HMI tags "DB_SDC_EMS"
   "SDC\DB_SDC_EMS\EMS[XXX].DISTANCE" : DInt AT %DB0.DBD0, 1 s   // Abstand zum vorangehenden EMS / distance to preciding EMS
   "SDC\DB_SDC_EMS\_Byte_EMS[XXX].ABS_POS" : Int, internal   // Absolute Position / absolute Positon
   "SDC\DB_SDC_EMS\EMS[XXX].IF_I_EMS.STAT" : DWord AT %DB0.DBD0, 1 s
   "SDC\DB_SDC_EMS\EMS[XXX].PRECEDING_EMS" : Int AT %DB0.DBW0, 1 s   // preciding EMS
   "SDC\DB_SDC_EMS\_Byte_EMS[XXX].TS_STAT.VAL.SEK" : Int, internal   // Sektion
   "SDC\DB_SDC_EMS\_Byte_EMS[XXX].DISTANCE" : Int, internal   // Abstand zum vorangehenden EMS / distance to preciding EMS
   "DB_SDC_EMS_HMI_HEADER.START_HMI" : Int = PLC DB_SDC_EMS_HMI.HEADER.START_HMI AT %DB3814.DBW16, 1 s   // Startadresse HMI
   "SDC\DB_SDC_EMS\EMS[XXX].IF_I_EMS.EA1" : DWord AT %DB0.DBD0, 1 s
   "SDC\DB_SDC_EMS\HMI[XX].PROFIL_Nr" : Int AT %DB0.DBW0, 1 s   // Profilnummer
   "SDC\DB_SDC_EMS\_EMS_HMI_Byte_16" : Int, internal
   "SDC\DB_SDC_EMS\HMI[XX].T_EDIT" : Bool AT %DB0.DBX0.0, 1 s   // Taster Editieren für Pult aktivieren
   "SDC\DB_SDC_EMS\_EMS_HMI_Byte_18" : Int, internal
   "SDC\DB_SDC_EMS\EMS[XXX].FKT_RESET" : Word AT %DB0.DBW0, 1 s   // EMS zur Reperatur / EMS to Repair
   "SDC\DB_SDC_EMS\EMS[XXX].IF_Q_EMS.D_SETSPEED" : DInt AT %DB0.DBD0, 1 s   // set value: drive speed (mm/min)
   "SDC\DB_SDC_EMS\_Byte_EMS[XXX].CYCLE_COUNTER" : Int, internal   // Zykluszähler / Cycle Counter
   "SDC\DB_SDC_EMS\HMI[XX].FR_EDIT" : Bool AT %DB0.DBX0.0, 1 s   // Freigabe Editieren
   "SDC\DB_SDC_EMS\_Byte_EMS[XXX].IF_I_EMS.H_POS" : Int, internal
   "SDC\DB_SDC_EMS\EMS[XXX].TS_STAT.SERIES" : Array [0..3] of Char AT %DB0.DBX0.0, 1 s   // Entwicklungs Serie Karosse (e.g. E-90, E-87 ) / Development series body (e.g. E-90, E-87 )
   "SDC\DB_SDC_EMS\EMS[XXX].IF_Q_EMS.D_SETPOS" : DInt AT %DB0.DBD0, 1 s   // Setpoint: drive position in mm
   "SDC\DB_SDC_EMS\HMI[XX].BILD_Nr_Alt" : Int AT %DB0.DBW0, 1 s   // Bild_Nr alt
   "SDC\DB_SDC_EMS\EMS[XXX].IF_Q_EMS.H_SETSPEED" : Int AT %DB0.DBW0, 1 s   // Setpoint: hoist speed (mm/min)
   "SDC\DB_SDC_EMS\_EMS_HMI_Byte_10" : Int, internal
   "SDC\DB_SDC_EMS\EMS[XXX].IF_I_EMS.H_POS" : Int AT %DB0.DBW0, 1 s
   "SDC\DB_SDC_EMS\_Byte_EMS[XXX].IF_Q_EMS.D_SETPOS" : Int, internal   // Setpoint: drive position in mm Pointer
   "SDC\DB_SDC_EMS\HMI[XX].EMS_Nr" : Int AT %DB0.DBW0, 1 s   // Sektionsnummer
   "SDC\DB_SDC_EMS\_Byte_EMS[XXX].PRECEDING_EMS" : Int, internal   // preciding EMS
   "SDC\DB_SDC_EMS\_Byte_EMS[XXX].IF_I_EMS.STAT" : Int, internal
   "SDC\DB_SDC_EMS\_EMS_HMI_Byte_09" : Int, internal
   "SDC\DB_SDC_EMS\_Byte_EMS[XXX].ERRORS_SDC" : Int, internal   // Fehler SDC Pointer / Faults SDC Pointer
   "SDC\DB_SDC_EMS\EMS[XXX].FLAGS" : Word AT %DB0.DBW0, 1 s   // EMS antrieb vorhanden / EMSdriver present
   "SDC\DB_SDC_EMS\_Byte_EMS[XXX].IF_I_EMS.EA2" : Int, internal
   "SDC\DB_SDC_EMS\EMS[XXX].ERRORS_SDC" : Word AT %DB0.DBW0, 1 s   // Fehler SDC / Faults SDC
   "SDC\DB_SDC_EMS\HMI[XX].T_SAVE" : Bool AT %DB0.DBX0.2, 1 s   // Taster speichern
   "SDC\DB_SDC_EMS\_Byte_EMS[XXX].PROFIL" : Int, internal   // Profile Number
   "SDC\DB_SDC_EMS\_Byte_EMS[XXX].FLAGS" : Int, internal   // EMS antrieb vorhanden / EMSdriver present
   "DB_SDC_EMS_1_HEADER.START_EMS" : Int = PLC DB_SDC_EMS_1.HEADER.START_EMS AT %DB3714.DBW6, 1 s   // Startadresse der EMS Daten im Daten DB
   "SDC\DB_SDC_EMS\EMS[XXX].IF_I_EMS.EA2" : DWord AT %DB0.DBD0, 1 s
   "SDC\DB_SDC_EMS\EMS[XXX].TS_STAT.VAL.SEK" : Int AT %DB0.DBW0, 1 s   // Sektion
      on ChangeValue: "SDC_TS_REFERENCE"("SDC\DB_SDC_EMS\EMS[XXX].TS_STAT.VAL.SEK")
   "SDC\DB_SDC_EMS\EMS[XXX].IF_I_EMS.D_POS" : DInt AT %DB0.DBD0, 1 s
   "SDC\DB_SDC_EMS\_Byte_EMS[XXX].IF_Q_EMS.H_SETSPEED" : Int, internal   // Setpoint: hoist speed (mm/min) Pointer
   "DB_SDC_EMS_1_HEADER.LAENGE_EMS" : Int = PLC DB_SDC_EMS_1.HEADER.LAENGE_EMS AT %DB3714.DBW8, 1 s   // Länge Eingänge pro EMS
   "SDC\DB_SDC_EMS\_EMS_HMI_Byte_19" : Int, internal
   "DB_SDC_EMS_1_HEADER.MIN_NR_EMS" : Int = PLC DB_SDC_EMS_1.HEADER.MIN_NR_EMS AT %DB3714.DBW2, 1 s   // Niedrigste EMS Nummer im Daten DB
   "SDC\DB_SDC_EMS\_Byte_EMS[XXX].IF_Q_EMS.H_SETPOS" : Int, internal   // Setpoint: hoist position (mm) Pointer
   "SDC\DB_SDC_EMS\_Byte_EMS[XXX].IF_I_EMS.EA1" : Int, internal
   "SDC\DB_SDC_EMS\_Intern_DB_EMS_Nr" : Int, internal
   "SDC\DB_SDC_EMS\HMI[XX].ER_DATA" : Bool AT %DB0.DBX0.1, 1 s   // Daten Fehlerhaft
   "DB_SDC_EMS_1_HEADER.OFFSET_EMS_FKT" : Int = PLC DB_SDC_EMS_1.HEADER.OFFSET_EMS_FKT AT %DB3714.DBW14, 1 s   // Offset EMS Funktions
   "SDC\DB_SDC_EMS\EMS[XXX].IF_Q_EMS.H_SETPOS" : Int AT %DB0.DBW0, 1 s   // Setpoint: hoist position (mm)
   "SDC\DB_SDC_EMS\_Byte_EMS[XXX].IF_I_EMS.ERROR" : Int, internal   // Fehlernummer Pointer / Error number Pointer
   "SDC\DB_SDC_EMS\_Byte_EMS[XXX].FKT_RESET" : Int, internal   // EMS zur Reperatur / EMS to Repair
   "SDC\DB_SDC_EMS\EMS[XXX].IF_Q_EMS.CONT" : DWord AT %DB0.DBD0, 1 s
   "DB_SDC_EMS_HMI_HEADER.OFFEST_HMI_DATA" : Int = PLC DB_SDC_EMS_HMI.HEADER.OFFEST_HMI_DATA AT %DB3814.DBW18, 1 s   // Offestadresse der HMI EMS Data
   "SDC\DB_SDC_EMS\_Byte_EMS[XXX].FKT_SET" : Int, internal   // EMS zur Reperatur / EMS to Repair
   "SDC\DB_SDC_EMS\HMI[XX].PULT_Nr_EDIT" : Int AT %DB0.DBW0, 1 s   // Pult Nr Editieren Aktiv (HMI 1 = Master)
   "SDC\DB_SDC_EMS\_EMS_HMI_Byte_00" : Int, internal
   "DB_SDC_EMS_1_HEADER.MAX_NR_EMS" : Int = PLC DB_SDC_EMS_1.HEADER.MAX_NR_EMS AT %DB3714.DBW4, 1 s   // Höchste EMS Nummer im Daten DB
   "SDC\DB_SDC_EMS\EMS[XXX].IF_I_EMS.ERROR" : Int AT %DB0.DBW0, 1 s   // Fehlernummer / Error number
   "DB_SDC_EMS_1_HEADER.OFFSET_EMS_SEK_STAT" : Int = PLC DB_SDC_EMS_1.HEADER.OFFSET_EMS_SEK_STAT AT %DB3714.DBW10, 1 s   // Offset EMS Data
   "DB_SDC_EMS_1_HEADER.LAENGE_EMS_SEK_STAT" : Int = PLC DB_SDC_EMS_1.HEADER.LAENGE_EMS_SEK_STAT AT %DB3714.DBW12, 1 s   // Länge EMS Data
   "SDC\DB_SDC_EMS\_Byte_EMS[XXX].TS_STAT.SERIES" : Int, internal   // Entwicklungs Serie Karosse (e.g. E-90, E-87 ) / Development series body (e.g. E-90, E-87 )
   "SDC\DB_SDC_EMS\HMI[XX].BILD_Nr" : Int AT %DB0.DBW0, 1 s   // Bild_Nr aktiv
   "SDC\DB_SDC_EMS\EMS[XXX].CYCLE_COUNTER" : Int AT %DB0.DBW0, 1 s   // Zykluszähler / Cycle Counter
   "SDC\DB_SDC_EMS\EMS[XXX].FKT_SET" : Word AT %DB0.DBW0, 1 s   // EMS zur Reperatur / EMS to Repair
      on ChangeValue: ResetBit("SDC\DB_SDC_EMS\_Intern_EMS_FKT_Info_Rep_1_on"); ResetBit("SDC\DB_SDC_EMS\_Intern_EMS_FKT_Info_Rep_2_on")
   "SDC\DB_SDC_EMS\HMI[XX].T_LOAD" : Bool AT %DB0.DBX0.3, 1 s   // Taster laden
   "SDC\DB_SDC_EMS\_EMS_HMI_Byte_12" : Int, internal
   "SDC\DB_SDC_EMS\_EMS_HMI_Byte_04" : Int, internal
   "DB_SDC_EMS_HMI_HMI[1].PULT_Nr_EDIT" : Int = PLC DB_SDC_EMS_HMI.HMI[1].PULT_Nr_EDIT AT %DB3814.DBW20, 1 s   // Pult Nr Editieren Aktiv (HMI 1 = Master)
   "SDC\DB_SDC_EMS\_EMS_HMI_Byte_14" : Int, internal
   "SDC\DB_SDC_EMS\_EMS_HMI_Byte_06" : Int, internal
   "SDC\DB_SDC_EMS\_Byte_EMS[XXX].IF_I_EMS.D_POS" : Int, internal
   "SDC\DB_SDC_EMS\_EMS_HMI_Byte_08" : Int, internal
   "SDC\DB_SDC_EMS\EMS[XXX].PROFIL" : Int AT %DB0.DBW0, 1 s   // Profile Number
      on ChangeValue: "SDC_GLOBAL_REFERENCE_PROFIL"("SDC\DB_SDC_EMS\EMS[XXX].PROFIL")
   "SDC\DB_SDC_EMS\_EMS_HMI_Byte_02" : Int, internal
   "SDC\DB_SDC_EMS\EMS[XXX].ABS_POS" : DInt AT %DB0.DBD0, 1 s   // absolute Positon
   "SDC\DB_SDC_EMS\HMI[XX].T_RESET_BED" : Bool AT %DB0.DBX0.1, 1 s   // Taster Reset Bedienfreigabe Pult Nr Bedienung
   "SDC\DB_SDC_EMS\_Byte_EMS[XXX].IF_Q_EMS.CONT" : Int, internal
   "SDC\DB_SDC_EMS\_Byte_EMS[XXX].IF_Q_EMS.D_SETSPEED" : Int, internal   // set value: drive speed (mm/min) Pointer
   "SDC\DB_SDC_EMS\_Byte_EMS[XXX].TS_STAT.VAL.ERROR" : Int, internal   // Sektion
   "SDC\DB_SDC_EMS\EMS[XXX].TS_STAT.VAL.ERROR" : Int AT %DB0.DBW0, 1 s   // Sektion
      on ChangeValue: SetTag("_DB_SDC_ERRORS.Error_nr", "SDC\DB_SDC_EMS\EMS[XXX].TS_STAT.VAL.ERROR")
   "DB_SDC_EMS_HMI_HEADER.DB_NR" : Int = PLC DB_SDC_EMS_HMI.HEADER.DB_NR AT %DB3814.DBW0, 1 s   // DB Nummer
   "SDC\DB_SDC_EMS\_Byte_EMS[XXX].IF_Q_EMS.T_SETPOS" : Int, internal   // Setpoint: hoist position (mm) Pointer
   "SDC\DB_SDC_EMS\_Byte_EMS[XXX].IF_Q_EMS.T_SETSPEED" : Int, internal   // Setpoint: hoist speed (mm/min) Pointer
   "SDC\DB_SDC_EMS\EMS[XXX].IF_Q_EMS.T_SETPOS" : Int AT %DB0.DBW0, 1 s   // Setpoint: hoist position (mm)
   "SDC\DB_SDC_EMS\EMS[XXX].IF_Q_EMS.T_SETSPEED" : Int AT %DB0.DBW0, 1 s   // Setpoint: hoist speed (mm/min)
   "SDC\DB_SDC_EMS\_Byte_EMS[XXX].IF_I_EMS.T_POS" : Int, internal
   "SDC\DB_SDC_EMS\EMS[XXX].IF_I_EMS.T_POS" : Int AT %DB0.DBW0, 1 s
   "SDC\DB_SDC_EMS\_Byte_EMS[XXX].FKT_INFO_REP_1" : Int, internal
   "SDC\DB_SDC_EMS\_Byte_EMS[XXX].FKT_INFO_REP_2" : Int, internal
   "SDC\DB_SDC_EMS\EMS[XXX].FKT_INFO_REP_1" : Int AT %DB0.DBW0, 1 s
   "SDC\DB_SDC_EMS\EMS[XXX].FKT_INFO_REP_2" : Int AT %DB0.DBW0, 1 s
   "SDC\DB_SDC_EMS\_Intern_EMS_FKT_Info_Rep_1_on" : Bool, internal
   "SDC\DB_SDC_EMS\_Intern_EMS_FKT_Info_Rep_2_on" : Bool, internal
   "SDC\DB_SDC_EMS\EMS[XXX].IF_I_EMS.EA3" : Word AT %DB0.DBW0, 1 s
   "SDC\DB_SDC_EMS\_Byte_EMS[XXX].IF_I_EMS.EA3" : Int, internal
   "SDC\DB_SDC_EMS\_Byte_EMS[XXX].VersNo[0]" : Int, internal   // Zykluszähler / Cycle Counter
   "SDC\DB_SDC_EMS\_Byte_EMS[XXX].VersNo[1]" : Int, internal   // Zykluszähler / Cycle Counter
   "SDC\DB_SDC_EMS\EMS[XXX].VersNo[0]" : Byte AT %DB0.DBB0, 1 s   // Zykluszähler / Cycle Counter
   "SDC\DB_SDC_EMS\EMS[XXX].VersNo[1]" : Byte AT %DB0.DBB0, 1 s   // Zykluszähler / Cycle Counter

HMI tags "DB_SDC_SIM"
   "DB_SDC_EMS_SIM_PAR.ON" : Bool = PLC DB_SDC_EMS_SIM.PAR.ON AT %DB3726.DBX40.0, 1 s   // Simulation ON "1"
   "DB_SDC_EMS_SIM_PAR.LEAP_AKT" : Array [0..19] of Bool = PLC DB_SDC_EMS_SIM.PAR.LEAP_AKT AT %DB3726.DBX32.0, 1 s   // Leap Aktiv
   "DB_SDC_EMS_SIM_PAR.BARCODE_START" : DInt = PLC DB_SDC_EMS_SIM.PAR.BARCODE_START AT %DB3726.DBD20, 1 s   // min Barcodevalue
   "DB_SDC_EMS_SIM_PAR.HUB_ENDE" : Int = PLC DB_SDC_EMS_SIM.PAR.HUB_ENDE AT %DB3726.DBW30, 1 s   // max Hoistvalue
   "DB_SDC_EMS_SIM_EMS[2].D_POS" : DInt = PLC DB_SDC_EMS_SIM.EMS[2].D_POS AT %DB3726.DBD90, 1 s   // Antriebsposition in mm / Drive position in mm
   "DB_SDC_EMS_SIM_PAR.BARCODE_ENDE" : DInt = PLC DB_SDC_EMS_SIM.PAR.BARCODE_ENDE AT %DB3726.DBD24, 1 s   // max Barcodevalue
   "DB_SDC_EMS_SIM_PAR.HUB_START" : Int = PLC DB_SDC_EMS_SIM.PAR.HUB_START AT %DB3726.DBW28, 1 s   // min Hoistvalue
   "DB_SDC_EMS_SIM_EMS[1].D_POS" : DInt = PLC DB_SDC_EMS_SIM.EMS[1].D_POS AT %DB3726.DBD50, 1 s   // Antriebsposition in mm / Drive position in mm
   "DB_SDC_EMS_SIM_EMS[3].D_POS" : DInt = PLC DB_SDC_EMS_SIM.EMS[3].D_POS AT %DB3726.DBD130, 1 s   // Antriebsposition in mm / Drive position in mm

HMI tags "DB_SDC_ERRORS"
   "DB_SDC_ERRORS_HEADER.DB_NR" : Int = PLC DB_SDC_ERRORS.HEADER.DB_NR AT %DB3722.DBW0, 1 s
   "DB_SDC_ERRORS_HEADER.MIN_NR_EMS" : Int = PLC DB_SDC_ERRORS.HEADER.MIN_NR_EMS AT %DB3722.DBW2, 1 s
   "DB_SDC_ERRORS_HEADER.MAX_NR_EMS" : Int = PLC DB_SDC_ERRORS.HEADER.MAX_NR_EMS AT %DB3722.DBW4, 1 s
   "DB_SDC_ERRORS_HEADER.START_EMS" : Int = PLC DB_SDC_ERRORS.HEADER.START_EMS AT %DB3722.DBW6, 1 s
   "DB_SDC_ERRORS_HEADER.LAENGE_EMS_StörungS" : Int = PLC DB_SDC_ERRORS.HEADER.LAENGE_EMS_StörungS AT %DB3722.DBW8, 1 s
   "DB_SDC_ERRORS.EMS[XXX].GEN_1" : Word AT %DB0.DBW0, 1 s
   "_Byte_DB_SDC_ERRORS.EMS[XXX].GEN_1" : UInt, internal
   "DB_SDC_ERRORS.EMS[XXX].GEN_2" : Word AT %DB0.DBW0, 1 s
   "_Byte_DB_SDC_ERRORS.EMS[XXX].GEN_2" : UInt, internal
   "DB_SDC_ERRORS.EMS[XXX].GEN_3" : Word AT %DB0.DBW0, 1 s
   "_Byte_DB_SDC_ERRORS.EMS[XXX].GEN_3" : UInt, internal
   "DB_SDC_ERRORS.EMS[XXX].GEN_4" : Word AT %DB0.DBW0, 1 s
   "_Byte_DB_SDC_ERRORS.EMS[XXX].GEN_4" : UInt, internal
   "DB_SDC_ERRORS.EMS[XXX].DRIVE_1" : Word AT %DB0.DBW0, 1 s
   "_Byte_DB_SDC_ERRORS.EMS[XXX].DRIVE_1" : UInt, internal
   "DB_SDC_ERRORS.EMS[XXX].DRIVE_2" : Word AT %DB0.DBW0, 1 s
   "_Byte_DB_SDC_ERRORS.EMS[XXX].DRIVE_2" : UInt, internal
   "DB_SDC_ERRORS.EMS[XXX].FC_DRIVE_1" : Word AT %DB0.DBW0, 1 s
   "_Byte_DB_SDC_ERRORS.EMS[XXX].FC_DRIVE_1" : UInt, internal
   "DB_SDC_ERRORS.EMS[XXX].FC_DRIVE_2" : Word AT %DB0.DBW0, 1 s
   "_Byte_DB_SDC_ERRORS.EMS[XXX].FC_DRIVE_2" : UInt, internal
   "DB_SDC_ERRORS.EMS[XXX].SAFETY_DRIVE" : Word AT %DB0.DBW0, 1 s
   "_Byte_DB_SDC_ERRORS.EMS[XXX].SAFETY_DRIVE" : UInt, internal
   "_Byte_DB_SDC_ERRORS.EMS[XXX].HOIST_1" : UInt, internal
   "DB_SDC_ERRORS.EMS[XXX].HOIST_2" : Word AT %DB0.DBW0, 1 s
   "_Byte_DB_SDC_ERRORS.EMS[XXX].HOIST_2" : UInt, internal
   "DB_SDC_ERRORS.EMS[XXX].FC_HOIST_1" : Word AT %DB0.DBW0, 1 s
   "_Byte_DB_SDC_ERRORS.EMS[XXX].FC_HOIST_1" : UInt, internal
   "DB_SDC_ERRORS.EMS[XXX].FC_HOIST_2" : Word AT %DB0.DBW0, 1 s
   "_Byte_DB_SDC_ERRORS.EMS[XXX].FC_HOIST_2" : UInt, internal
   "DB_SDC_ERRORS.EMS[XXX].SAFETY_HOIST" : Word AT %DB0.DBW0, 1 s
   "_Byte_DB_SDC_ERRORS.EMS[XXX].SAFETY_HOIST" : UInt, internal
   "DB_SDC_ERRORS.EMS[XXX].HOIST_1" : Word AT %DB0.DBW0, 1 s
   "_Byte_DB_SDC_ERRORS.EMS[XXX].TILT_1" : UInt, internal
   "DB_SDC_ERRORS.EMS[XXX].TILT_2" : Word AT %DB0.DBW0, 1 s
   "_Byte_DB_SDC_ERRORS.EMS[XXX].TILT_2" : UInt, internal
   "DB_SDC_ERRORS.EMS[XXX].FC_TILT_1" : Word AT %DB0.DBW0, 1 s
   "_Byte_DB_SDC_ERRORS.EMS[XXX].FC_TILT_1" : UInt, internal
   "DB_SDC_ERRORS.EMS[XXX].FC_TILT_2" : Word AT %DB0.DBW0, 1 s
   "_Byte_DB_SDC_ERRORS.EMS[XXX].FC_TILT_2" : UInt, internal
   "DB_SDC_ERRORS.EMS[XXX].SAFETY_TILT" : Word AT %DB0.DBW0, 1 s
   "_Byte_DB_SDC_ERRORS.EMS[XXX].SAFETY_TILT" : UInt, internal
   "DB_SDC_ERRORS.EMS[XXX].TILT_1" : Word AT %DB0.DBW0, 1 s
   "DB_SDC_ERRORS.EMS[XXX].SDC" : Word AT %DB0.DBW0, 1 s
   "_Byte_DB_SDC_ERRORS.EMS[XXX].SDC" : UInt, internal
   "DB_SDC_ERRORS.SDC" : Word AT %DB3722.DBW20020, 1 s
   "_DB_SDC_ERRORS.Error_nr" : Int, internal

HMI tags "DB_SDC_GLOBAL_REFERENCE"
   "DB_SDC_GLOBAL_REFERENCE_PAR_SET[8].LIMITS" : Array [0..15] of Char = PLC DB_SDC_GLOBAL_REFERENCE.PAR_SET[8].LIMITS AT %DB3786.DBX292.0, 1 s
   "DB_SDC_GLOBAL_REFERENCE_PAR_SET[3].LIMITS" : Array [0..15] of Char = PLC DB_SDC_GLOBAL_REFERENCE.PAR_SET[3].LIMITS AT %DB3786.DBX132.0, 1 s
   "DB_SDC_GLOBAL_REFERENCE_PAR_SET[0].LIMITS" : Array [0..15] of Char = PLC DB_SDC_GLOBAL_REFERENCE.PAR_SET[0].LIMITS AT %DB3786.DBX36.0, 1 s
   "DB_SDC_GLOBAL_REFERENCE_PAR_SET[14].SYNCH" : Array [0..15] of Char = PLC DB_SDC_GLOBAL_REFERENCE.PAR_SET[14].SYNCH AT %DB3786.DBX468.0, 1 s
   "DB_SDC_GLOBAL_REFERENCE_PAR_SET[9].SYNCH" : Array [0..15] of Char = PLC DB_SDC_GLOBAL_REFERENCE.PAR_SET[9].SYNCH AT %DB3786.DBX308.0, 1 s
   "DB_SDC_GLOBAL_REFERENCE_PAR_SET[11].LIMITS" : Array [0..15] of Char = PLC DB_SDC_GLOBAL_REFERENCE.PAR_SET[11].LIMITS AT %DB3786.DBX388.0, 1 s
   "DB_SDC_GLOBAL_REFERENCE_PAR_SET[10].LIMITS" : Array [0..15] of Char = PLC DB_SDC_GLOBAL_REFERENCE.PAR_SET[10].LIMITS AT %DB3786.DBX356.0, 1 s
   "DB_SDC_GLOBAL_REFERENCE_PAR_SET[0].SYNCH" : Array [0..15] of Char = PLC DB_SDC_GLOBAL_REFERENCE.PAR_SET[0].SYNCH AT %DB3786.DBX20.0, 1 s
   "DB_SDC_GLOBAL_REFERENCE_PAR_SET[14].LIMITS" : Array [0..15] of Char = PLC DB_SDC_GLOBAL_REFERENCE.PAR_SET[14].LIMITS AT %DB3786.DBX484.0, 1 s
   "DB_SDC_GLOBAL_REFERENCE_PAR_SET[6].LIMITS" : Array [0..15] of Char = PLC DB_SDC_GLOBAL_REFERENCE.PAR_SET[6].LIMITS AT %DB3786.DBX228.0, 1 s
   "DB_SDC_GLOBAL_REFERENCE_PAR_SET[10].SYNCH" : Array [0..15] of Char = PLC DB_SDC_GLOBAL_REFERENCE.PAR_SET[10].SYNCH AT %DB3786.DBX340.0, 1 s
   "DB_SDC_GLOBAL_REFERENCE_PAR_SET[5].SYNCH" : Array [0..15] of Char = PLC DB_SDC_GLOBAL_REFERENCE.PAR_SET[5].SYNCH AT %DB3786.DBX180.0, 1 s
   "DB_SDC_GLOBAL_REFERENCE_PAR_SET[13].SYNCH" : Array [0..15] of Char = PLC DB_SDC_GLOBAL_REFERENCE.PAR_SET[13].SYNCH AT %DB3786.DBX436.0, 1 s
   "DB_SDC_GLOBAL_REFERENCE_PAR_SET[12].LIMITS" : Array [0..15] of Char = PLC DB_SDC_GLOBAL_REFERENCE.PAR_SET[12].LIMITS AT %DB3786.DBX420.0, 1 s
   "DB_SDC_GLOBAL_REFERENCE_PAR_SET[15].SYNCH" : Array [0..15] of Char = PLC DB_SDC_GLOBAL_REFERENCE.PAR_SET[15].SYNCH AT %DB3786.DBX500.0, 1 s
   "DB_SDC_GLOBAL_REFERENCE_PAR_SET[2].LIMITS" : Array [0..15] of Char = PLC DB_SDC_GLOBAL_REFERENCE.PAR_SET[2].LIMITS AT %DB3786.DBX100.0, 1 s
   "DB_SDC_GLOBAL_REFERENCE_PAR_SET[6].SYNCH" : Array [0..15] of Char = PLC DB_SDC_GLOBAL_REFERENCE.PAR_SET[6].SYNCH AT %DB3786.DBX212.0, 1 s
   "DB_SDC_GLOBAL_REFERENCE_PAR_SET[1].SYNCH" : Array [0..15] of Char = PLC DB_SDC_GLOBAL_REFERENCE.PAR_SET[1].SYNCH AT %DB3786.DBX52.0, 1 s
   "DB_SDC_GLOBAL_REFERENCE_PAR_SET[4].SYNCH" : Array [0..15] of Char = PLC DB_SDC_GLOBAL_REFERENCE.PAR_SET[4].SYNCH AT %DB3786.DBX148.0, 1 s
   "DB_SDC_GLOBAL_REFERENCE_PAR_SET[8].SYNCH" : Array [0..15] of Char = PLC DB_SDC_GLOBAL_REFERENCE.PAR_SET[8].SYNCH AT %DB3786.DBX276.0, 1 s
   "DB_SDC_GLOBAL_REFERENCE_PAR_SET[2].SYNCH" : Array [0..15] of Char = PLC DB_SDC_GLOBAL_REFERENCE.PAR_SET[2].SYNCH AT %DB3786.DBX84.0, 1 s
   "DB_SDC_GLOBAL_REFERENCE_PAR_SET[1].LIMITS" : Array [0..15] of Char = PLC DB_SDC_GLOBAL_REFERENCE.PAR_SET[1].LIMITS AT %DB3786.DBX68.0, 1 s
   "DB_SDC_GLOBAL_REFERENCE_PAR_SET[15].LIMITS" : Array [0..15] of Char = PLC DB_SDC_GLOBAL_REFERENCE.PAR_SET[15].LIMITS AT %DB3786.DBX516.0, 1 s
   "DB_SDC_GLOBAL_REFERENCE_PAR_SET[11].SYNCH" : Array [0..15] of Char = PLC DB_SDC_GLOBAL_REFERENCE.PAR_SET[11].SYNCH AT %DB3786.DBX372.0, 1 s
   "DB_SDC_GLOBAL_REFERENCE_PAR_SET[3].SYNCH" : Array [0..15] of Char = PLC DB_SDC_GLOBAL_REFERENCE.PAR_SET[3].SYNCH AT %DB3786.DBX116.0, 1 s
   "DB_SDC_GLOBAL_REFERENCE_PAR_SET[4].LIMITS" : Array [0..15] of Char = PLC DB_SDC_GLOBAL_REFERENCE.PAR_SET[4].LIMITS AT %DB3786.DBX164.0, 1 s
   "DB_SDC_GLOBAL_REFERENCE_PAR_SET[12].SYNCH" : Array [0..15] of Char = PLC DB_SDC_GLOBAL_REFERENCE.PAR_SET[12].SYNCH AT %DB3786.DBX404.0, 1 s
   "DB_SDC_GLOBAL_REFERENCE_PAR_SET[9].LIMITS" : Array [0..15] of Char = PLC DB_SDC_GLOBAL_REFERENCE.PAR_SET[9].LIMITS AT %DB3786.DBX324.0, 1 s
   "DB_SDC_GLOBAL_REFERENCE_PAR_SET[7].SYNCH" : Array [0..15] of Char = PLC DB_SDC_GLOBAL_REFERENCE.PAR_SET[7].SYNCH AT %DB3786.DBX244.0, 1 s
   "DB_SDC_GLOBAL_REFERENCE_PAR_SET[7].LIMITS" : Array [0..15] of Char = PLC DB_SDC_GLOBAL_REFERENCE.PAR_SET[7].LIMITS AT %DB3786.DBX260.0, 1 s
   "DB_SDC_GLOBAL_REFERENCE_PAR_SET[13].LIMITS" : Array [0..15] of Char = PLC DB_SDC_GLOBAL_REFERENCE.PAR_SET[13].LIMITS AT %DB3786.DBX452.0, 1 s
   "DB_SDC_GLOBAL_REFERENCE_PAR_SET[5].LIMITS" : Array [0..15] of Char = PLC DB_SDC_GLOBAL_REFERENCE.PAR_SET[5].LIMITS AT %DB3786.DBX196.0, 1 s
   "SDC\DB_SDC_GLOBAL_REFERENCE\DB_SDC_GLOBAL_REFERENCE.PROFIL[XX].SORTE" : Array [0..5] of Char AT %DB0.DBX0.0, 1 s
   "DB_SDC_GLOBAL_REFERENCE_HEADER.START_PROFIL" : Int = PLC DB_SDC_GLOBAL_REFERENCE.HEADER.START_PROFIL AT %DB3786.DBW14, 1 s
   "DB_SDC_GLOBAL_REFERENCE_HEADER.LAENGE_PROFIL" : Int = PLC DB_SDC_GLOBAL_REFERENCE.HEADER.LAENGE_PROFIL AT %DB3786.DBW16, 1 s
   "_DB_SDC_GLOBAL_REFERENCE.PROFIL[XX].SORTE_Byte" : Int, internal
   "DB_SDC_GLOBAL_REFERENCE_HEADER.MIN_PROFIL" : Int = PLC DB_SDC_GLOBAL_REFERENCE.HEADER.MIN_PROFIL AT %DB3786.DBW10, 1 s
   "DB_SDC_GLOBAL_REFERENCE_HEADER.MAX_PROFIL" : Int = PLC DB_SDC_GLOBAL_REFERENCE.HEADER.MAX_PROFIL AT %DB3786.DBW12, 1 s
   "_DB_SDC_GLOBAL_REFERENCE.PROFIL[XX+1].SORTE_Byte" : Int, internal
   "SDC\DB_SDC_GLOBAL_REFERENCE\DB_SDC_GLOBAL_REFERENCE.PROFIL[XX+1].SORTE" : Array [0..5] of Char AT %DB0.DBX0.0, 1 s
   "DB_SDC_GLOBAL_REFERENCE_HEADER.DB_NR" : Int = PLC DB_SDC_GLOBAL_REFERENCE.HEADER.DB_NR AT %DB3786.DBW0, 1 s

HMI tags "DB_SDC_EMS_TA"
   "DB_SDC_EMS_TA_HEADER.DB_NR" : Int = PLC DB_SDC_EMS_TA.HEADER.DB_NR AT %DB3728.DBW0, 1 s
   "DB_SDC_EMS_TA_HEADER.MIN_NR_EMS" : Int = PLC DB_SDC_EMS_TA.HEADER.MIN_NR_EMS AT %DB3728.DBW2, 1 s
   "DB_SDC_EMS_TA_HEADER.MAX_NR_EMS" : Int = PLC DB_SDC_EMS_TA.HEADER.MAX_NR_EMS AT %DB3728.DBW4, 1 s
   "DB_SDC_EMS_TA_HEADER.START_EMS" : Int = PLC DB_SDC_EMS_TA.HEADER.START_EMS AT %DB3728.DBW6, 1 s
   "DB_SDC_EMS_TA_HEADER.LAENGE_TA_DATA" : Int = PLC DB_SDC_EMS_TA.HEADER.LAENGE_TA_DATA AT %DB3728.DBW8, 1 s
   "DB_SDC_EMS_TA_HEADER.ANZ_TA" : Int = PLC DB_SDC_EMS_TA.HEADER.ANZ_TA AT %DB3728.DBW10, 1 s
   "DB_SDC_EMS_TA.EMS[XX].TA1.PW1" : Int AT %DB0.DBW0, 1 s
   "_Byte_DB_SDC_EMS_TA.EMS[XX].TA1.PW1" : DInt, internal
   "_Byte_DB_SDC_EMS_TA.EMS[XX].TA1.PW2" : DInt, internal
   "_Byte_DB_SDC_EMS_TA.EMS[XX].TA1.PW3" : DInt, internal
   "_Byte_DB_SDC_EMS_TA.EMS[XX].TA2.PW1" : DInt, internal
   "_Byte_DB_SDC_EMS_TA.EMS[XX].TA2.PW2" : DInt, internal
   "_Byte_DB_SDC_EMS_TA.EMS[XX].TA2.PW3" : DInt, internal
   "_Byte_DB_SDC_EMS_TA.EMS[XX].TA3.PW1" : DInt, internal
   "_Byte_DB_SDC_EMS_TA.EMS[XX].TA3.PW2" : DInt, internal
   "_Byte_DB_SDC_EMS_TA.EMS[XX].TA3.PW3" : DInt, internal
   "DB_SDC_EMS_TA.EMS[XX].TA1.PW2" : Int AT %DB0.DBW0, 1 s
   "DB_SDC_EMS_TA.EMS[XX].TA1.PW3" : Int AT %DB0.DBW0, 1 s
   "DB_SDC_EMS_TA.EMS[XX].TA2.PW1" : Int AT %DB0.DBW0, 1 s
   "DB_SDC_EMS_TA.EMS[XX].TA2.PW2" : Int AT %DB0.DBW0, 1 s
   "DB_SDC_EMS_TA.EMS[XX].TA2.PW3" : Int AT %DB0.DBW0, 1 s
   "DB_SDC_EMS_TA.EMS[XX].TA3.PW1" : Int AT %DB0.DBW0, 1 s
   "DB_SDC_EMS_TA.EMS[XX].TA3.PW2" : Int AT %DB0.DBW0, 1 s
   "DB_SDC_EMS_TA.EMS[XX].TA3.PW3" : Int AT %DB0.DBW0, 1 s
   "DB_SDC_EMS_TA.EMS[XX].TA1.FAULT" : Int AT %DB0.DBW0, 1 s
   "_Byte_DB_SDC_EMS_TA.EMS[XX].TA1.FAULT" : Int AT %MW36, 1 s
   "_Byte_DB_SDC_EMS_TA.EMS[XX].TA1.ALARM" : Int AT %MW38, 1 s
   "_Byte_DB_SDC_EMS_TA.EMS[XX].TA2.FAULT" : DInt, internal
   "_Byte_DB_SDC_EMS_TA.EMS[XX].TA2.ALARM" : DInt, internal
   "_Byte_DB_SDC_EMS_TA.EMS[XX].TA3.FAULT" : DInt, internal
   "_Byte_DB_SDC_EMS_TA.EMS[XX].TA3.ALARM" : DInt, internal
   "DB_SDC_EMS_TA.EMS[XX].TA1.ALARM" : Int AT %DB0.DBW0, 1 s

HMI tags "DB_SDC_TS_IF"
   "DB_SDC_TS_IF_COMMAND_HEADER.DB_NR" : Int = PLC DB_SDC_TS_IF_COMMAND.HEADER.DB_NR AT %DB3716.DBW0, 1 s
   "DB_SDC_TS_IF_COMMAND_HEADER.MIN_NR_SEK" : Int = PLC DB_SDC_TS_IF_COMMAND.HEADER.MIN_NR_SEK AT %DB3716.DBW2, 1 s
   "DB_SDC_TS_IF_COMMAND_HEADER.MAX_NR_SEK" : Int = PLC DB_SDC_TS_IF_COMMAND.HEADER.MAX_NR_SEK AT %DB3716.DBW4, 1 s
   "DB_SDC_TS_IF_COMMAND_HEADER.START_DAT" : Int = PLC DB_SDC_TS_IF_COMMAND.HEADER.START_DAT AT %DB3716.DBW6, 1 s
   "DB_SDC_TS_IF_COMMAND_HEADER.LAENGE_SEK_DATA" : Int = PLC DB_SDC_TS_IF_COMMAND.HEADER.LAENGE_SEK_DATA AT %DB3716.DBW8, 1 s
   "DB_SDC_TS_IF_COMMAND.SEK[XXX].VAL.PROFIL" : Int AT %DB0.DBW0, 1 s
   "_Byte_DB_SDC_TS_IF_COMMAND.SEK[XXX].VAL.PROFIL" : Int, internal
   "DB_SDC_TS_IF_COMMAND_2_HEADER.DB_NR" : Int = PLC DB_SDC_TS_IF_COMMAND_2.HEADER.DB_NR AT %DB3717.DBW0, 1 s
   "DB_SDC_TS_IF_COMMAND_2_HEADER.LAENGE_SEK_DATA" : Int = PLC DB_SDC_TS_IF_COMMAND_2.HEADER.LAENGE_SEK_DATA AT %DB3717.DBW8, 1 s
   "DB_SDC_TS_IF_COMMAND_2_HEADER.MAX_NR_SEK" : Int = PLC DB_SDC_TS_IF_COMMAND_2.HEADER.MAX_NR_SEK AT %DB3717.DBW4, 1 s
   "DB_SDC_TS_IF_COMMAND_2_HEADER.MIN_NR_SEK" : Int = PLC DB_SDC_TS_IF_COMMAND_2.HEADER.MIN_NR_SEK AT %DB3717.DBW2, 1 s
   "DB_SDC_TS_IF_COMMAND_2_HEADER.START_DAT" : Int = PLC DB_SDC_TS_IF_COMMAND_2.HEADER.START_DAT AT %DB3717.DBW6, 1 s
   "_DB_SDC_TS_IF_COMMAND.HEADER.DB_NR" : Int AT %DB716.DBW0
   "_Byte_DB_SDC_TS_IF_COMMAND.SEK[XXX].VAL.D_SETSPEED" : Int, internal
   "DB_SDC_TS_IF_COMMAND.SEK[XXX].VAL.D_SETSPEED" : DInt AT %DB0.DBD0, 1 s
   "_Byte_DB_SDC_TS_IF_COMMAND.SEK[XXX].VAL.D_POS_OFFS" : Int, internal
   "DB_SDC_TS_IF_COMMAND.SEK[XXX].VAL.D_POS_OFFS" : Int AT %DB0.DBW0, 1 s
   "_Byte_DB_SDC_TS_IF_COMMAND.SEK[XXX].BIT1" : Int, internal
   "DB_SDC_TS_IF_COMMAND.SEK[XXX].BIT1" : Int AT %DB0.DBW0, 1 s
   "DB_SDC_TS_IF_COMMAND.SEK[XXX].BIT2" : Int AT %DB0.DBW0, 1 s
   "_Byte_DB_SDC_TS_IF_COMMAND.SEK[XXX].BIT2" : Int, internal
   "DB_SDC_TS_IF_COMMAND.SEK[XXX].BIT3" : Int AT %DB0.DBW0, 1 s
   "_Byte_DB_SDC_TS_IF_COMMAND.SEK[XXX].BIT3" : Int, internal
   "DB_SDC_TS_IF_COMMAND.SEK[XXX].FKT_SET" : Int AT %DB0.DBW0, 1 s
   "_Byte_DB_SDC_TS_IF_COMMAND.SEK[XXX].FKT_SET" : Int, internal
   "DB_SDC_TS_IF_COMMAND.SEK[XXX].FKT_RESET" : Int AT %DB0.DBW0, 1 s
   "_Byte_DB_SDC_TS_IF_COMMAND.SEK[XXX].FKT_RESET" : Int, internal
   "_DB_SDC_TS_IF_STATUS.HEADER.DB_NR" : Int AT %DB716.DBW0
   "_Byte_DB_SDC_TS_IF_STATUS.SEK[XXX].BIT1" : Int, internal
   "_Byte_DB_SDC_TS_IF_STATUS.SEK[XXX].BIT2" : Int, internal
   "_Byte_DB_SDC_TS_IF_STATUS.SEK[XXX].BIT3" : Int, internal
   "_Byte_DB_SDC_TS_IF_STATUS.SEK[XXX].FKT_SET" : Int, internal
   "_Byte_DB_SDC_TS_IF_STATUS.SEK[XXX].VAL.DRIVE_POS" : Int, internal
   "_Byte_DB_SDC_TS_IF_STATUS.SEK[XXX].VAL.PROFIL" : Int, internal
   "_Byte_DB_SDC_TS_IF_STATUS.SEK[XXX].VAL.EMS_ID" : Int, internal
   "DB_SDC_TS_IF_STATUS_HEADER.DB_NR" : Int = PLC DB_SDC_TS_IF_STATUS.HEADER.DB_NR AT %DB3718.DBW0, 1 s
   "DB_SDC_TS_IF_STATUS_HEADER.LAENGE_SEK_DATA" : Int = PLC DB_SDC_TS_IF_STATUS.HEADER.LAENGE_SEK_DATA AT %DB3718.DBW8, 1 s
   "DB_SDC_TS_IF_STATUS_HEADER.MAX_NR_SEK" : Int = PLC DB_SDC_TS_IF_STATUS.HEADER.MAX_NR_SEK AT %DB3718.DBW4, 1 s
   "DB_SDC_TS_IF_STATUS_HEADER.MIN_NR_SEK" : Int = PLC DB_SDC_TS_IF_STATUS.HEADER.MIN_NR_SEK AT %DB3718.DBW2, 1 s
   "DB_SDC_TS_IF_STATUS_HEADER.START_DAT" : Int = PLC DB_SDC_TS_IF_STATUS.HEADER.START_DAT AT %DB3718.DBW6, 1 s
   "DB_SDC_TS_IF_STATUS.SEK[XXX].BIT1" : Int AT %DB0.DBW0, 1 s
   "DB_SDC_TS_IF_STATUS.SEK[XXX].BIT2" : Int AT %DB0.DBW0, 1 s
   "DB_SDC_TS_IF_STATUS.SEK[XXX].BIT3" : Int AT %DB0.DBW0, 1 s
   "DB_SDC_TS_IF_STATUS.SEK[XXX].FKT_SET" : Int AT %DB0.DBW0, 1 s
   "DB_SDC_TS_IF_STATUS.SEK[XXX].VAL.DRIVE_POS" : DInt AT %DB0.DBD0, 1 s
   "DB_SDC_TS_IF_STATUS.SEK[XXX].VAL.PROFIL" : Int AT %DB0.DBW0, 1 s
   "DB_SDC_TS_IF_STATUS.SEK[XXX].VAL.EMS_ID" : Int AT %DB0.DBW0, 1 s
   "DB_SDC_TS_IF_STATUS_2_HEADER.DB_NR" : Int = PLC DB_SDC_TS_IF_STATUS_2.HEADER.DB_NR AT %DB3719.DBW0, 1 s
   "DB_SDC_TS_IF_STATUS_2_HEADER.LAENGE_SEK_DATA" : Int = PLC DB_SDC_TS_IF_STATUS_2.HEADER.LAENGE_SEK_DATA AT %DB3719.DBW8, 1 s
   "DB_SDC_TS_IF_STATUS_2_HEADER.MAX_NR_SEK" : Int = PLC DB_SDC_TS_IF_STATUS_2.HEADER.MAX_NR_SEK AT %DB3719.DBW4, 1 s
   "DB_SDC_TS_IF_STATUS_2_HEADER.MIN_NR_SEK" : Int = PLC DB_SDC_TS_IF_STATUS_2.HEADER.MIN_NR_SEK AT %DB3719.DBW2, 1 s
   "DB_SDC_TS_IF_STATUS_2_HEADER.START_DAT" : Int = PLC DB_SDC_TS_IF_STATUS_2.HEADER.START_DAT AT %DB3719.DBW6, 1 s
   "DB_SDC_TS_IF_STATUS.SEK[XXX].BIT4" : Int AT %DB0.DBW0, 1 s
   "_Byte_DB_SDC_TS_IF_STATUS.SEK[XXX].BIT4" : Int, internal
   "DB_SDC_TS_IF_STATUS.SEK[XXX].SORTE" : Array [0..3] of Char AT %DB0.DBX0.0, 1 s
   "_Byte_DB_SDC_TS_IF_STATUS.SEK[XXX].SORTE" : Int, internal
   "DB_SDC_TS_IF_STATUS.SEK[XXX].VAL.HOIST_POS" : Int AT %DB0.DBW0, 1 s
   "_Byte_DB_SDC_TS_IF_STATUS.SEK[XXX].VAL.HOIST_POS" : Int, internal
   "DB_SDC_TS_IF_STATUS.SEK[XXX].VAL.TILT_POS" : Int AT %DB0.DBW0, 1 s
   "_Byte_DB_SDC_TS_IF_STATUS.SEK[XXX].VAL.TILT_POS" : Int, internal
   "DB_SDC_TS_IF_STATUS.SEK[XXX].VAL.ERROR" : Int AT %DB0.DBW0, 1 s
   "_Byte_DB_SDC_TS_IF_STATUS.SEK[XXX].VAL.ERROR" : Int, internal
   "DB_SDC_TS_IF_STATUS.SEK[XXX].VAL.DRIVE_POS_PERC" : Int AT %DB0.DBW0, 1 s
   "_Byte_DB_SDC_TS_IF_STATUS.SEK[XXX].VAL.DRIVE_POS_PERC" : Int, internal
   "DB_SDC_TS_IF_STATUS.SEK[XXX].VAL.SEK" : Int AT %DB0.DBW0, 1 s
   "_Byte_DB_SDC_TS_IF_STATUS.SEK[XXX].VAL.SEK" : Int, internal
   "DB_SDC_TS_IF_HMI_HEADER.DB_NR" : Int = PLC DB_SDC_TS_IF_HMI.HEADER.DB_NR AT %DB3816.DBW0, 1 s
   "DB_SDC_TS_IF_HMI_HEADER.START_DAT" : Int = PLC DB_SDC_TS_IF_HMI.HEADER.START_DAT AT %DB3816.DBW6, 1 s
   "DB_SDC_TS_IF_HMI_HEADER.LAENGE_SEK_COM" : Int = PLC DB_SDC_TS_IF_HMI.HEADER.LAENGE_SEK_COM AT %DB3816.DBW8, 1 s
   "DB_SDC_TS_IF_HMI_HEADER.LAENGE_SEK_STAT" : Int = PLC DB_SDC_TS_IF_HMI.HEADER.LAENGE_SEK_STAT AT %DB3816.DBW10, 1 s
   "DB_SDC_TS_IF_HMI_HEADER.OFFEST_SEK_STAT" : Int = PLC DB_SDC_TS_IF_HMI.HEADER.OFFEST_SEK_STAT AT %DB3816.DBW12, 1 s
   "DB_SDC_TS_IF_HMI_HEADER.START_HMI" : Int = PLC DB_SDC_TS_IF_HMI.HEADER.START_HMI AT %DB3816.DBW16, 1 s
   "DB_SDC_TS_IF_HMI_HEADER.OFFEST_HMI_DATA" : Int = PLC DB_SDC_TS_IF_HMI.HEADER.OFFEST_HMI_DATA AT %DB3816.DBW18, 1 s
   "_DB_SDC_TS_IF_HMI.HMI_Byte_00" : Int, internal
   "_DB_SDC_TS_IF_HMI.HMI_Byte_02" : Int, internal
   "_DB_SDC_TS_IF_HMI.HMI_Byte_04" : Int, internal
   "_DB_SDC_TS_IF_HMI.HMI_Byte_06" : Int, internal
   "_DB_SDC_TS_IF_HMI.HMI_Byte_08" : Int, internal
   "_DB_SDC_TS_IF_HMI.HMI_Byte_09" : Int, internal
   "_DB_SDC_TS_IF_HMI.HMI_Byte_10" : Int, internal
   "_DB_SDC_TS_IF_HMI.HMI_Byte_12" : Int, internal
   "_DB_SDC_TS_IF_HMI.HMI_Byte_14" : Int, internal
   "_DB_SDC_TS_IF_HMI.HMI_Byte_16" : Int, internal
   "_DB_SDC_TS_IF_HMI.HMI_Byte_18" : Int, internal
   "_DB_SDC_TS_IF_HMI.HMI_Byte_19" : Int, internal
   "DB_SDC_TS_IF_HMI.HMI[XX].BILD_Nr" : Int AT %DB0.DBW0, 1 s   // Bild_Nr aktiv
   "DB_SDC_TS_IF_HMI.HMI[XX].SEK_Nr" : Int AT %DB0.DBW0, 1 s   // Bild_Nr aktiv

HMI tags "DB_SDC_EMS_PAR_ALLG"
   "DB_SDC_EMS_PAR_HMI_HEADER.DB_NR" : Int = PLC DB_SDC_EMS_PAR_HMI.HEADER.DB_NR AT %DB3802.DBW0, 1 s
   "DB_SDC_EMS_PAR_HMI_HEADER.START_PAR" : Int = PLC DB_SDC_EMS_PAR_HMI.HEADER.START_PAR AT %DB3802.DBW6, 1 s
   "DB_SDC_EMS_PAR_HMI_HEADER.LAENGE_PAR" : Int = PLC DB_SDC_EMS_PAR_HMI.HEADER.LAENGE_PAR AT %DB3802.DBW8, 1 s
   "DB_SDC_EMS_PAR_HMI_HMI[1].PULT_Nr_EDIT" : Int = PLC DB_SDC_EMS_PAR_HMI.HMI[1].PULT_Nr_EDIT AT %DB3802.DBW20, 1 s
   "DB_SDC_EMS_PAR_HMI.HMI[XX].BILD_Nr" : Int AT %DB0.DBW0, 1 s
   "DB_SDC_EMS_PAR_HMI.HMI[XX].BILD_Nr_Alt" : Int AT %DB0.DBW0, 1 s
   "_PAR_HMI_Byte_00" : Int, internal
   "_PAR_HMI_Byte_02" : Int, internal
   "_PAR_HMI_Byte_04" : Int, internal
   "_PAR_HMI_Byte_06" : Int, internal
   "_PAR_HMI_Byte_08" : Int, internal
   "_PAR_HMI_Byte_09" : Int, internal
   "_PAR_HMI_Byte_10" : Int, internal
   "_PAR_HMI_Byte_12" : Int, internal
   "_PAR_HMI_Byte_14" : Int, internal
   "_PAR_HMI_Byte_16" : Int, internal
   "_PAR_HMI_Byte_18" : Int, internal
   "_PAR_HMI_Byte_19" : Int, internal
   "DB_SDC_EMS_PAR_HMI.HMI[XX].FR_EDIT" : Bool AT %DB0.DBX0.0, 1 s   // Freigabe Editieren
   "DB_SDC_EMS_PAR_HMI.HMI[XX].PULT_Nr_EDIT" : Int AT %DB0.DBW0, 1 s   // Pult Nr Editieren Aktiv (HMI 1 = Master)
   "DB_SDC_EMS_PAR_HMI.HMI[XX].T_EDIT" : Bool AT %DB0.DBX0.0, 1 s   // Taster Editieren für Pult aktivieren
   "DB_SDC_EMS_PAR_HMI.HMI[XX].T_LOAD" : Bool AT %DB0.DBX0.3, 1 s   // Taster laden
   "DB_SDC_EMS_PAR_HMI.HMI[XX].T_RESET_BED" : Bool AT %DB0.DBX0.1, 1 s   // Taster Reset Bedienfreigabe Pult Nr Bedienung
   "DB_SDC_EMS_PAR_HMI.HMI[XX].T_SAVE" : Bool AT %DB0.DBX0.2, 1 s   // Taster speichern
   "DB_SDC_EMS_PAR_HMI.HMI[XX].ER_DATA" : Bool AT %DB0.DBX0.1, 1 s   // Freigabe Editieren
   "DB_SDC_EMS_PAR_HMI_HEADER.START_HMI" : Int = PLC DB_SDC_EMS_PAR_HMI.HEADER.START_HMI AT %DB3802.DBW16, 1 s
   "DB_SDC_EMS_PAR_HMI_HEADER.OFFEST_HMI_DATA" : Int = PLC DB_SDC_EMS_PAR_HMI.HEADER.OFFEST_HMI_DATA AT %DB3802.DBW18, 1 s
